
REGION Network 14
   RUNG wire#powerrail
      "FC111_HMI_Status"()
   END_RUNG
   // the same network as SCL:
   "FC111_HMI_Status"();
END_REGION

REGION Network 15
   RUNG wire#powerrail
      "FC500_FAULTS"()
   END_RUNG
   // the same network as SCL:
   "FC500_FAULTS"();
END_REGION

REGION Network 16
   RUNG wire#powerrail
      "FC502_FAULTS C11-C20"()
   END_RUNG
   // the same network as SCL:
   "FC502_FAULTS C11-C20"();
END_REGION

REGION Network 17
   RUNG wire#powerrail
      "FC503_FAULTS C21-C30"()
   END_RUNG
   // the same network as SCL:
   "FC503_FAULTS C21-C30"();
END_REGION

REGION Network 18
   RUNG wire#powerrail
      "FC504_FAULTS C31-C40"()
   END_RUNG
   // the same network as SCL:
   "FC504_FAULTS C31-C40"();
END_REGION

REGION Network 19
   RUNG wire#powerrail
      "FC505_FAULTS C41-C50"()
   END_RUNG
   // the same network as SCL:
   "FC505_FAULTS C41-C50"();
END_REGION

REGION Network 20
   RUNG wire#powerrail
      "FC506_FAULTS C51-C60"()
   END_RUNG
   // the same network as SCL:
   "FC506_FAULTS C51-C60"();
END_REGION

REGION Network 21
   RUNG wire#powerrail
      "FC507_FAULTS C61-C70"()
   END_RUNG
   // the same network as SCL:
   "FC507_FAULTS C61-C70"();
END_REGION

REGION Network 22
   RUNG wire#powerrail
      "FC508_FAULTS C71-C80"()
   END_RUNG
   // the same network as SCL:
   "FC508_FAULTS C71-C80"();
END_REGION

REGION Network 23
   RUNG wire#powerrail
      "FC509_FAULTS C81-C82"()
   END_RUNG
   // the same network as SCL:
   "FC509_FAULTS C81-C82"();
END_REGION

REGION Network 24
   RUNG wire#powerrail
      "FC201_SDC_To_Carrier_Map_IO [C01-C10]"()
   END_RUNG
   // the same network as SCL:
   "FC201_SDC_To_Carrier_Map_IO [C01-C10]"();
END_REGION

REGION Network 25
   RUNG wire#powerrail
      "FC202_SDC_To_Carrier_Map_IO [C11-C20]"()
   END_RUNG
   // the same network as SCL:
   "FC202_SDC_To_Carrier_Map_IO [C11-C20]"();
END_REGION

REGION Network 26
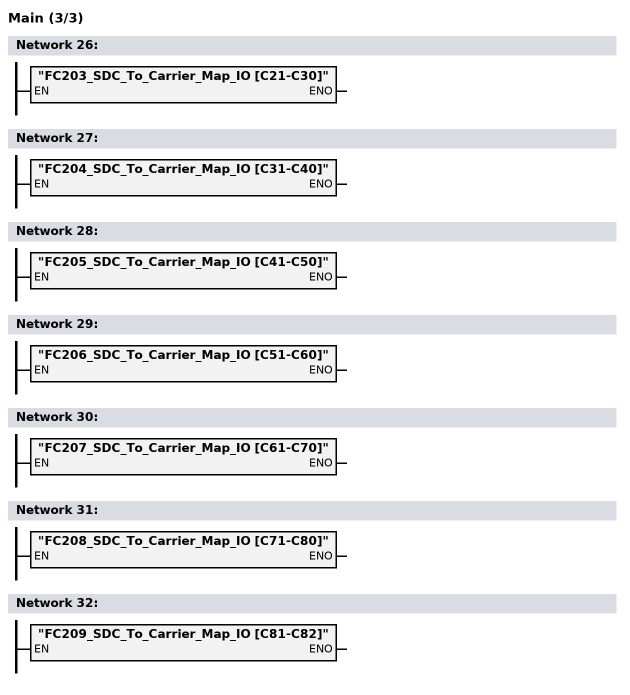
   RUNG wire#powerrail
      "FC203_SDC_To_Carrier_Map_IO [C21-C30]"()
   END_RUNG
   // the same network as SCL:
   "FC203_SDC_To_Carrier_Map_IO [C21-C30]"();
END_REGION

REGION Network 27
   RUNG wire#powerrail
      "FC204_SDC_To_Carrier_Map_IO [C31-C40]"()
   END_RUNG
   // the same network as SCL:
   "FC204_SDC_To_Carrier_Map_IO [C31-C40]"();
END_REGION

REGION Network 28
   RUNG wire#powerrail
      "FC205_SDC_To_Carrier_Map_IO [C41-C50]"()
   END_RUNG
   // the same network as SCL:
   "FC205_SDC_To_Carrier_Map_IO [C41-C50]"();
END_REGION

REGION Network 29
   RUNG wire#powerrail
      "FC206_SDC_To_Carrier_Map_IO [C51-C60]"()
   END_RUNG
   // the same network as SCL:
   "FC206_SDC_To_Carrier_Map_IO [C51-C60]"();
END_REGION

REGION Network 30
   RUNG wire#powerrail
      "FC207_SDC_To_Carrier_Map_IO [C61-C70]"()
   END_RUNG
   // the same network as SCL:
   "FC207_SDC_To_Carrier_Map_IO [C61-C70]"();
END_REGION

REGION Network 31
   RUNG wire#powerrail
      "FC208_SDC_To_Carrier_Map_IO [C71-C80]"()
   END_RUNG
   // the same network as SCL:
   "FC208_SDC_To_Carrier_Map_IO [C71-C80]"();
END_REGION

REGION Network 32
   RUNG wire#powerrail
      "FC209_SDC_To_Carrier_Map_IO [C81-C82]"()
   END_RUNG
   // the same network as SCL:
   "FC209_SDC_To_Carrier_Map_IO [C81-C82]"();
END_REGION
END_ORGANIZATION_BLOCK

ORGANIZATION_BLOCK "Startup"   // OB100, LAD, Startup
TITLE = "Complete Restart"
{ S7_Optimized_Access := 'TRUE' }
VERSION : 0.1
// //============================================================================
// //SIEMENS AG
// //(c)Copyright 2017 All Rights Reserved
// //-----------------------------------------------------------------------------
// //Library: -
// //Tested with: S7-1516-3 PN/DP FW 2.5
// //Engineering: TIA Portal V14 Update1
// //Restrictions: -
// //Requirements: -
// //Functionality: Startup OB for Diagnostics
// //-----------------------------------------------------------------------------
// //Change log table:
// //Version  Date              Expert in charge                               Changes applied
// //01.00.00 25.04.2017 Siemens Industry Online Support First released version
// //============================================================================
   VAR_INPUT
      LostRetentive : Bool;   // True if retentive data are lost
      LostRTC : Bool;   // True if date and time are lost
   END_VAR
   VAR_TEMP
      index : Int;
   END_VAR
BEGIN

REGION Network 1: Set start user diagnostic
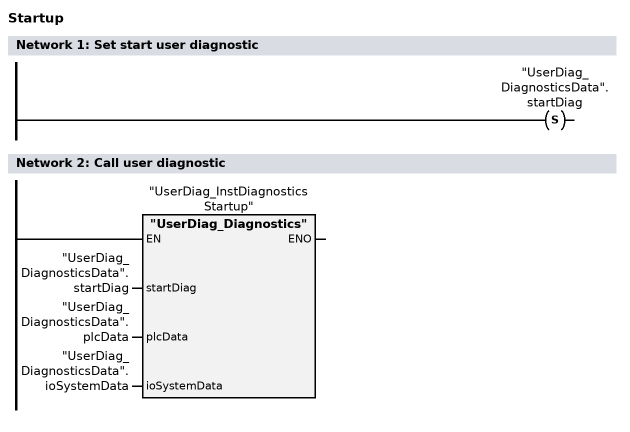
   RUNG wire#powerrail
      S_Coil( "UserDiag_DiagnosticsData".startDiag )
   END_RUNG
   // the same network as SCL:
   "UserDiag_DiagnosticsData".startDiag := TRUE;
END_REGION

REGION Network 2: Call user diagnostic
   RUNG wire#powerrail
      "UserDiag_InstDiagnosticsStartup"(startDiag := "UserDiag_DiagnosticsData".startDiag, plcData := "UserDiag_DiagnosticsData".plcData, ioSystemData := "UserDiag_DiagnosticsData".ioSystemData)
   END_RUNG
   // the same network as SCL:
   "UserDiag_InstDiagnosticsStartup"(startDiag := "UserDiag_DiagnosticsData".startDiag,   // "UserDiag_Diagnostics"
                           plcData := "UserDiag_DiagnosticsData".plcData,
                           ioSystemData := "UserDiag_DiagnosticsData".ioSystemData);
END_REGION
END_ORGANIZATION_BLOCK

ORGANIZATION_BLOCK "Cyclic SDC TO EMS"   // OB300, LAD, CyclicInterrupt
{ S7_Optimized_Access := 'TRUE' }
VERSION : 0.1
   VAR_INPUT
      Initial_Call : Bool;   // Initial call of this OB
      Event_Count : Int;   // Events discarded
   END_VAR
BEGIN
END_ORGANIZATION_BLOCK

// folder: 03_FBs

FUNCTION_BLOCK "FB110_FirstCarrierTCopMotionFB"   // FB110, LAD
{ S7_Optimized_Access := 'TRUE' }
VERSION : 0.1
   VAR_INPUT
      Zone : Int;
      ZonePos : Int;
      ClearOfStopDist : Int;
      StopControlFromEMS01 : "UDT_StopControlFromEMS01";
   END_VAR
   VAR_OUTPUT
      CarrierNumber : Int;
      MoveFwdCommand : Bool;
      DriveCmdSpeed : Int;
      NextCarrierNum : Word;
      NextStopPosition : DWord;
      AtCmdPosition : Bool;
      CarrierInTransitToNextZone : Bool;
      StopStatusToEMS01 : "UDT_StopStatusToEMS01";
   END_VAR
   VAR
      PreviousCarrierNumMemory : Word;
      TrafficCopCarrierZnBuffer : Array[0..40] of "UDT_TrafficCop";
      LastCarrierNextZnPos : Int;
      CarNumZnPos : Int;
      NextZone : Int;
      EndPos_LowLimit : DWord;
      EndPos_HighLimit : DWord;
      ClrOfStopPos_LowLimit : DWord;
      ClrOfStopPos_HighLimit : DWord;
      ClearOfStopPos : DWord;
      ClearToMoveTrain : Bool;
      PrevZone : Int;
      PrevZone_CarrierReady : Bool;
      LastCarrierCurrentZnPos : Int;
      LastCarrierNumber : Word;
      CarrierInTransitToProdZone : Bool;
      ResetCarrierInTransToProd : Bool;
      WaitPositionMemory : DInt;
      OneShot : Bool;
      NextCarrierOffset : DWord;
      PrevZone_EndPos_LowLimit : DWord;
      PrevZone_EndPos_HighLimit : DWord;
   END_VAR
   VAR_TEMP
      NextZoneBuffer : Int;
      LastZone : Int;
      HighSpeedSetpoint : Word;
      LowSpeedSetpoint : Word;
      NextZonePosition : Int;
      NextCarrierOffsetSetup1 : UDInt;
      NextCarrierOffsetSetup2 : UDInt;
   END_VAR
   VAR_TEMP   // added for the SCL form of the ladder/FBD networks
      _w1 : Bool;
      _w2 : Bool;
      _w3 : Bool;
      _w4 : Bool;
      _w5 : Bool;
   END_VAR
BEGIN

REGION Network 1
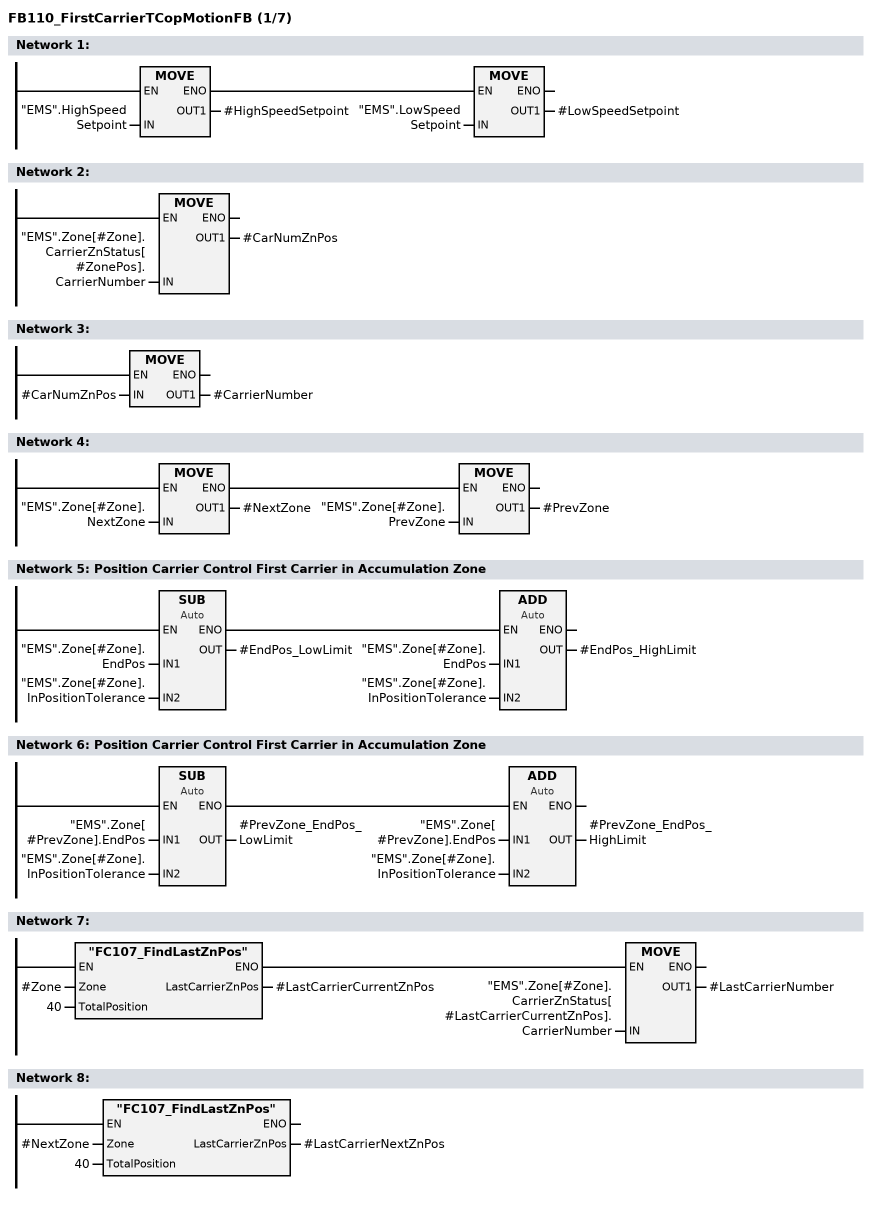
   RUNG wire#powerrail
      Move(in := "EMS".HighSpeedSetpoint, out1 => #HighSpeedSetpoint)
      Move(in := "EMS".LowSpeedSetpoint, out1 => #LowSpeedSetpoint)
   END_RUNG
   // the same network as SCL:
   #HighSpeedSetpoint := "EMS".HighSpeedSetpoint;
   #LowSpeedSetpoint := "EMS".LowSpeedSetpoint;
END_REGION

REGION Network 2
   RUNG wire#powerrail
      Move(in := "EMS".Zone[#Zone].CarrierZnStatus[#ZonePos].CarrierNumber, out1 => #CarNumZnPos)
   END_RUNG
   // the same network as SCL:
   #CarNumZnPos := "EMS".Zone[#Zone].CarrierZnStatus[#ZonePos].CarrierNumber;
END_REGION

REGION Network 3
   RUNG wire#powerrail
      Move(in := #CarNumZnPos, out1 => #CarrierNumber)
   END_RUNG
   // the same network as SCL:
   #CarrierNumber := #CarNumZnPos;
END_REGION

REGION Network 4
   RUNG wire#powerrail
      Move(in := "EMS".Zone[#Zone].NextZone, out1 => #NextZone)
      Move(in := "EMS".Zone[#Zone].PrevZone, out1 => #PrevZone)
   END_RUNG
   // the same network as SCL:
   #NextZone := "EMS".Zone[#Zone].NextZone;
   #PrevZone := "EMS".Zone[#Zone].PrevZone;
END_REGION

REGION Network 5: Position Carrier Control First Carrier in Accumulation Zone
   RUNG wire#powerrail
      Sub(in1 := "EMS".Zone[#Zone].EndPos, in2 := "EMS".Zone[#Zone].InPositionTolerance, out => #EndPos_LowLimit)
      Add(in1 := "EMS".Zone[#Zone].EndPos, in2 := "EMS".Zone[#Zone].InPositionTolerance, out => #EndPos_HighLimit)
   END_RUNG
   // the same network as SCL:
   #EndPos_LowLimit := "EMS".Zone[#Zone].EndPos - "EMS".Zone[#Zone].InPositionTolerance;
   #EndPos_HighLimit := "EMS".Zone[#Zone].EndPos + "EMS".Zone[#Zone].InPositionTolerance;
END_REGION

REGION Network 6: Position Carrier Control First Carrier in Accumulation Zone
   RUNG wire#powerrail
      Sub(in1 := "EMS".Zone[#PrevZone].EndPos, in2 := "EMS".Zone[#Zone].InPositionTolerance, out => #PrevZone_EndPos_LowLimit)
      Add(in1 := "EMS".Zone[#PrevZone].EndPos, in2 := "EMS".Zone[#Zone].InPositionTolerance, out => #PrevZone_EndPos_HighLimit)
   END_RUNG
   // the same network as SCL:
   #PrevZone_EndPos_LowLimit := "EMS".Zone[#PrevZone].EndPos - "EMS".Zone[#Zone].InPositionTolerance;
   #PrevZone_EndPos_HighLimit := "EMS".Zone[#PrevZone].EndPos + "EMS".Zone[#Zone].InPositionTolerance;
END_REGION

REGION Network 7
   RUNG wire#powerrail
      "FC107_FindLastZnPos"(Zone := #Zone, TotalPosition := 40, LastCarrierZnPos => #LastCarrierCurrentZnPos)
      Move(in := "EMS".Zone[#Zone].CarrierZnStatus[#LastCarrierCurrentZnPos].CarrierNumber, out1 => #LastCarrierNumber)
   END_RUNG
   // the same network as SCL:
   "FC107_FindLastZnPos"(Zone := #Zone,
                         TotalPosition := 40,
                         LastCarrierZnPos => #LastCarrierCurrentZnPos,
                         ENO => #_w1);
   IF #_w1 THEN
       #LastCarrierNumber := "EMS".Zone[#Zone].CarrierZnStatus[#LastCarrierCurrentZnPos].CarrierNumber;
   END_IF;
END_REGION

REGION Network 8
   RUNG wire#powerrail
      "FC107_FindLastZnPos"(Zone := #NextZone, TotalPosition := 40, LastCarrierZnPos => #LastCarrierNextZnPos)
   END_RUNG
   // the same network as SCL:
   "FC107_FindLastZnPos"(Zone := #NextZone, TotalPosition := 40, LastCarrierZnPos => #LastCarrierNextZnPos);
END_REGION

REGION Network 9: Position Carrier Control First Carrier in Production Zone
   // Control of First Carrier in Zone Closest to end position/Stop.  Move command is issued to carrier. Carrier will move in auto.
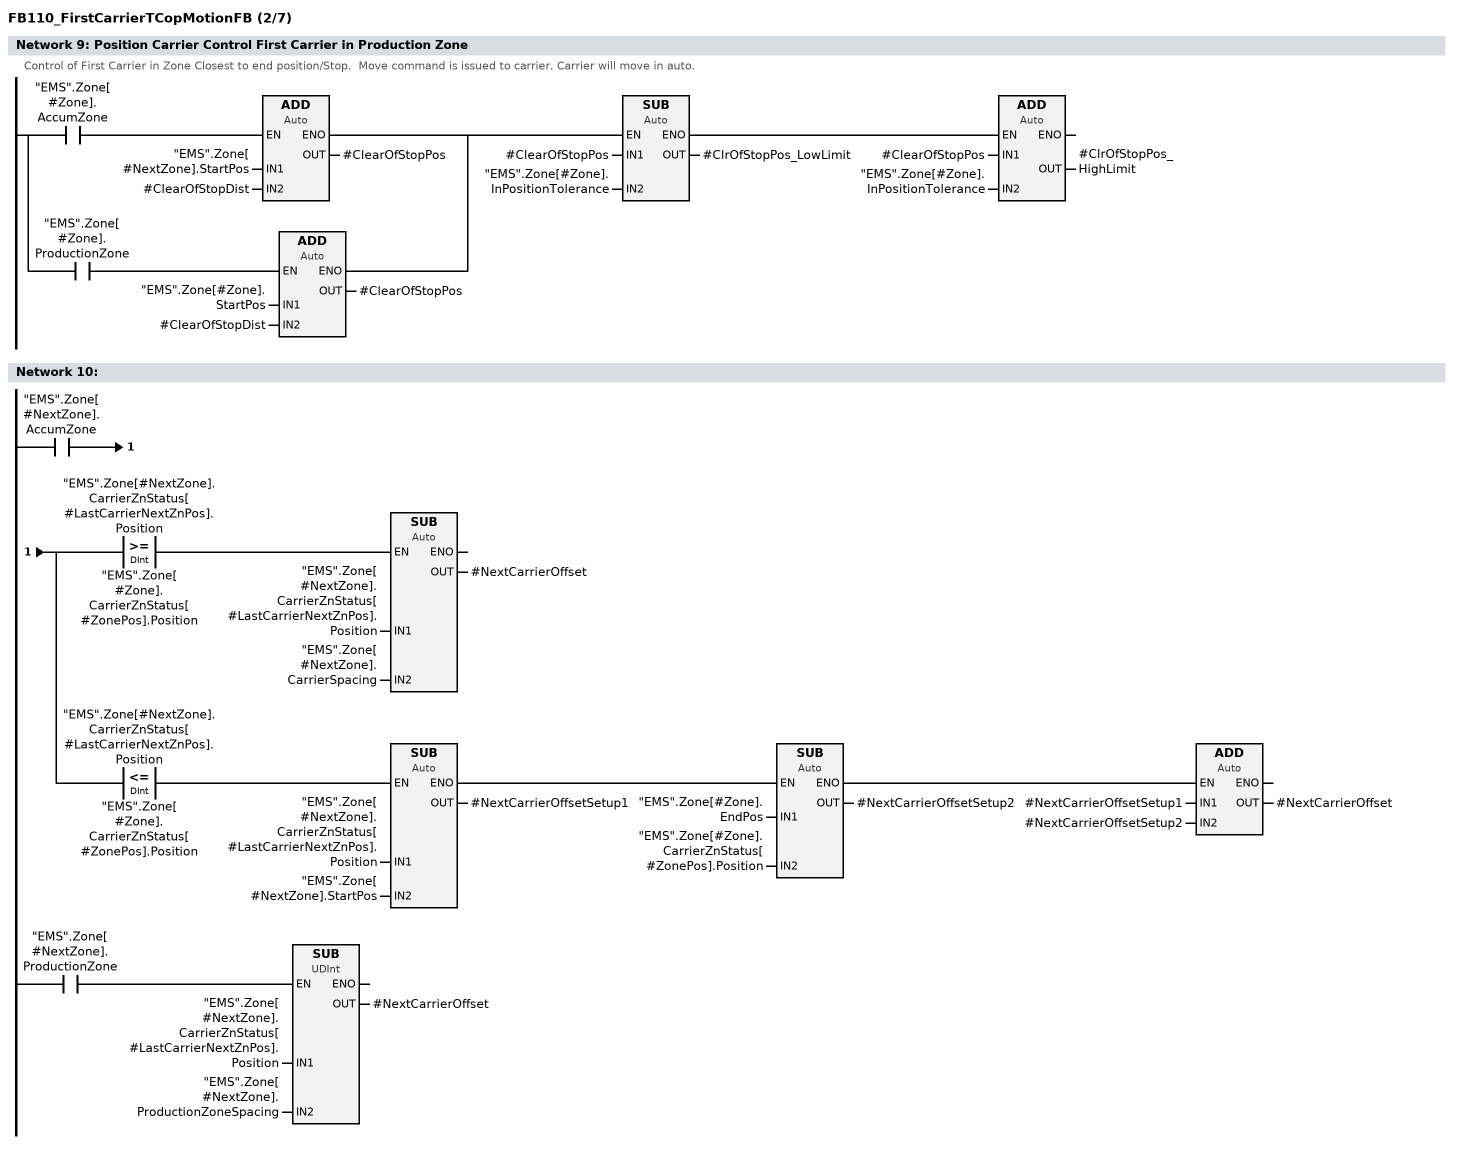
   RUNG wire#powerrail
      Contact( "EMS".Zone[#Zone].AccumZone )
      Add(in1 := "EMS".Zone[#NextZone].StartPos, in2 := #ClearOfStopDist, out => #ClearOfStopPos)
      wire#w1
      Sub(in1 := #ClearOfStopPos, in2 := "EMS".Zone[#Zone].InPositionTolerance, out => #ClrOfStopPos_LowLimit)
      Add(in1 := #ClearOfStopPos, in2 := "EMS".Zone[#Zone].InPositionTolerance, out => #ClrOfStopPos_HighLimit)
   END_RUNG
   RUNG wire#powerrail
      Contact( "EMS".Zone[#Zone].ProductionZone )
      Add(in1 := "EMS".Zone[#Zone].StartPos, in2 := #ClearOfStopDist, out => #ClearOfStopPos)
   END_RUNG wire#w1
   // the same network as SCL:
   IF "EMS".Zone[#Zone].AccumZone THEN
       #ClearOfStopPos := "EMS".Zone[#NextZone].StartPos + #ClearOfStopDist;
   END_IF;
   IF "EMS".Zone[#Zone].ProductionZone THEN
       #ClearOfStopPos := "EMS".Zone[#Zone].StartPos + #ClearOfStopDist;
   END_IF;
   IF "EMS".Zone[#Zone].AccumZone OR "EMS".Zone[#Zone].ProductionZone THEN
       #ClrOfStopPos_LowLimit := #ClearOfStopPos - "EMS".Zone[#Zone].InPositionTolerance;
       #ClrOfStopPos_HighLimit := #ClearOfStopPos + "EMS".Zone[#Zone].InPositionTolerance;
   END_IF;
END_REGION

REGION Network 10
   RUNG wire#powerrail
      Contact( "EMS".Zone[#NextZone].AccumZone )
      wire#w1
      { S7_Templates := "SrcType := DInt" } GE_Contact(in1 := "EMS".Zone[#NextZone].CarrierZnStatus[#LastCarrierNextZnPos].Position, in2 := "EMS".Zone[#Zone].CarrierZnStatus[#ZonePos].Position)
      Sub(in1 := "EMS".Zone[#NextZone].CarrierZnStatus[#LastCarrierNextZnPos].Position, in2 := "EMS".Zone[#NextZone].CarrierSpacing, out => #NextCarrierOffset)
   END_RUNG
   RUNG wire#w1
      { S7_Templates := "SrcType := DInt" } LE_Contact(in1 := "EMS".Zone[#NextZone].CarrierZnStatus[#LastCarrierNextZnPos].Position, in2 := "EMS".Zone[#Zone].CarrierZnStatus[#ZonePos].Position)
      Sub(in1 := "EMS".Zone[#NextZone].CarrierZnStatus[#LastCarrierNextZnPos].Position, in2 := "EMS".Zone[#NextZone].StartPos, out => #NextCarrierOffsetSetup1)
      Sub(in1 := "EMS".Zone[#Zone].EndPos, in2 := "EMS".Zone[#Zone].CarrierZnStatus[#ZonePos].Position, out => #NextCarrierOffsetSetup2)
      Add(in1 := #NextCarrierOffsetSetup1, in2 := #NextCarrierOffsetSetup2, out => #NextCarrierOffset)
   END_RUNG
   RUNG wire#powerrail
      Contact( "EMS".Zone[#NextZone].ProductionZone )
      { S7_Templates := "SrcType := UDInt" } Sub(in1 := "EMS".Zone[#NextZone].CarrierZnStatus[#LastCarrierNextZnPos].Position, in2 := "EMS".Zone[#NextZone].ProductionZoneSpacing, out => #NextCarrierOffset)
   END_RUNG
   // the same network as SCL:
   IF "EMS".Zone[#NextZone].AccumZone AND ("EMS".Zone[#NextZone].CarrierZnStatus[#LastCarrierNextZnPos].Position >= "EMS".Zone[#Zone].CarrierZnStatus[#ZonePos].Position) THEN
       #NextCarrierOffset := "EMS".Zone[#NextZone].CarrierZnStatus[#LastCarrierNextZnPos].Position - "EMS".Zone[#NextZone].CarrierSpacing;
   END_IF;
   IF "EMS".Zone[#NextZone].AccumZone AND ("EMS".Zone[#NextZone].CarrierZnStatus[#LastCarrierNextZnPos].Position <= "EMS".Zone[#Zone].CarrierZnStatus[#ZonePos].Position) THEN
       #NextCarrierOffsetSetup1 := "EMS".Zone[#NextZone].CarrierZnStatus[#LastCarrierNextZnPos].Position - "EMS".Zone[#NextZone].StartPos;
       #NextCarrierOffsetSetup2 := "EMS".Zone[#Zone].EndPos - "EMS".Zone[#Zone].CarrierZnStatus[#ZonePos].Position;
       #NextCarrierOffset := #NextCarrierOffsetSetup1 + #NextCarrierOffsetSetup2;
   END_IF;
   IF "EMS".Zone[#NextZone].ProductionZone THEN
       #NextCarrierOffset := "EMS".Zone[#NextZone].CarrierZnStatus[#LastCarrierNextZnPos].Position - "EMS".Zone[#NextZone].ProductionZoneSpacing;
   END_IF;
END_REGION

REGION Network 11
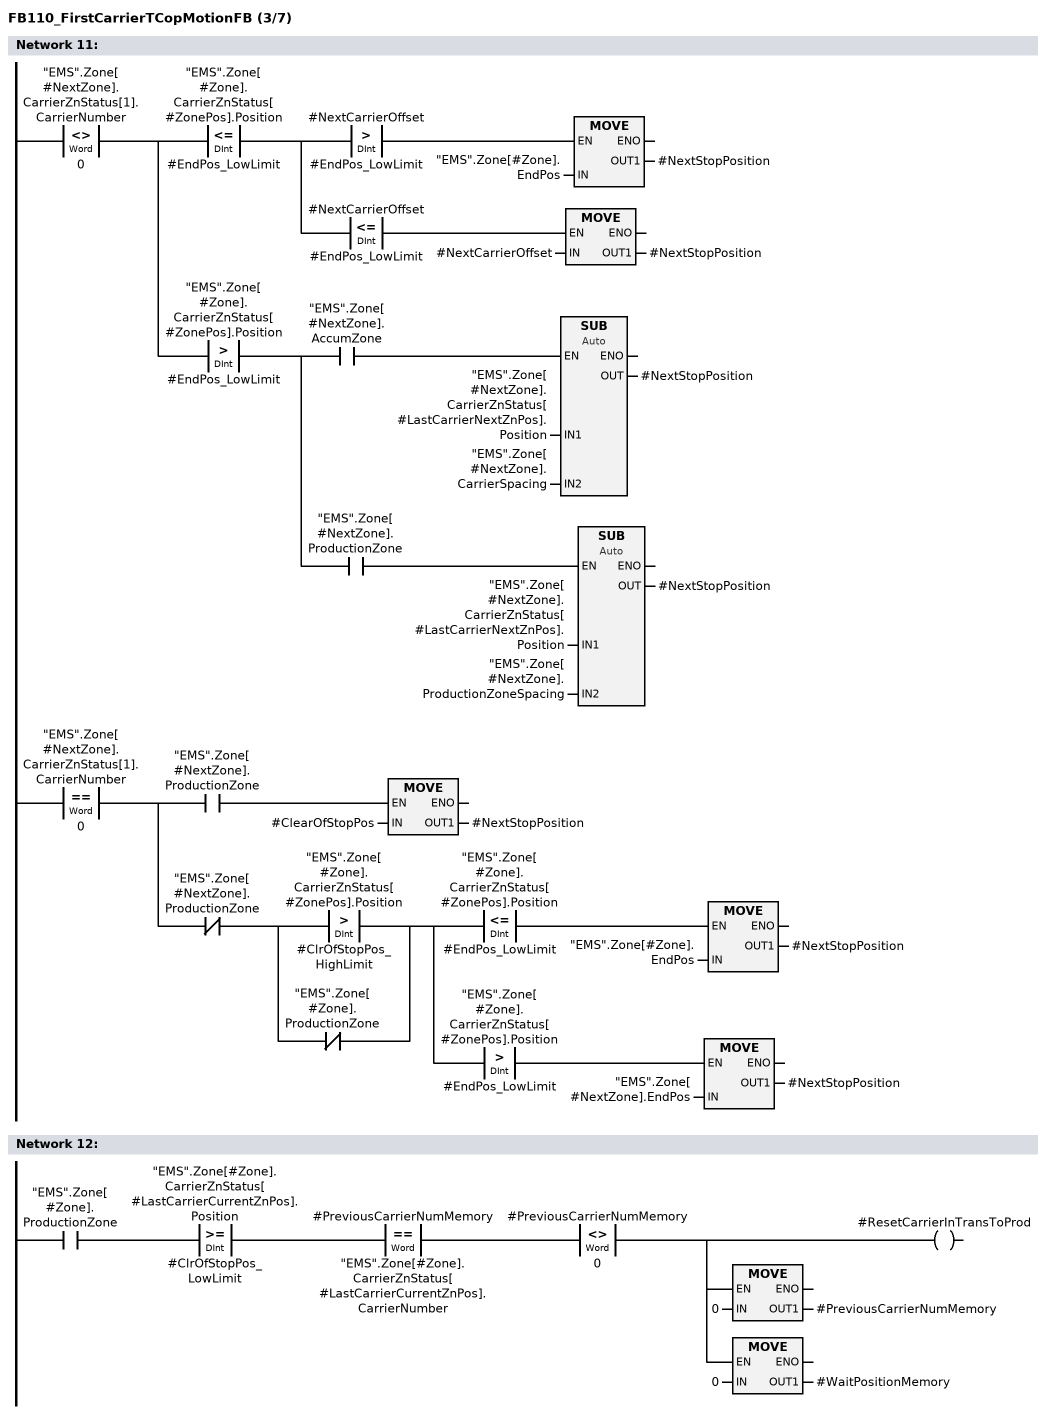
   RUNG wire#powerrail
      { S7_Templates := "SrcType := Word" } NE_Contact(in1 := "EMS".Zone[#NextZone].CarrierZnStatus[1].CarrierNumber, in2 := 0)
      wire#w1
      { S7_Templates := "SrcType := DInt" } LE_Contact(in1 := "EMS".Zone[#Zone].CarrierZnStatus[#ZonePos].Position, in2 := #EndPos_LowLimit)
      wire#w2
      { S7_Templates := "SrcType := DInt" } GT_Contact(in1 := #NextCarrierOffset, in2 := #EndPos_LowLimit)
      Move(in := "EMS".Zone[#Zone].EndPos, out1 => #NextStopPosition)
   END_RUNG
   RUNG wire#w2
      { S7_Templates := "SrcType := DInt" } LE_Contact(in1 := #NextCarrierOffset, in2 := #EndPos_LowLimit)
      Move(in := #NextCarrierOffset, out1 => #NextStopPosition)
   END_RUNG
   RUNG wire#w1
      { S7_Templates := "SrcType := DInt" } GT_Contact(in1 := "EMS".Zone[#Zone].CarrierZnStatus[#ZonePos].Position, in2 := #EndPos_LowLimit)
      wire#w3
      Contact( "EMS".Zone[#NextZone].AccumZone )
      Sub(in1 := "EMS".Zone[#NextZone].CarrierZnStatus[#LastCarrierNextZnPos].Position, in2 := "EMS".Zone[#NextZone].CarrierSpacing, out => #NextStopPosition)
   END_RUNG
   RUNG wire#w3
      Contact( "EMS".Zone[#NextZone].ProductionZone )
      Sub(in1 := "EMS".Zone[#NextZone].CarrierZnStatus[#LastCarrierNextZnPos].Position, in2 := "EMS".Zone[#NextZone].ProductionZoneSpacing, out => #NextStopPosition)
   END_RUNG
   RUNG wire#powerrail
      { S7_Templates := "SrcType := Word" } EQ_Contact(in1 := "EMS".Zone[#NextZone].CarrierZnStatus[1].CarrierNumber, in2 := 0)
      wire#w4
      Contact( "EMS".Zone[#NextZone].ProductionZone )
      Move(in := #ClearOfStopPos, out1 => #NextStopPosition)
   END_RUNG
   RUNG wire#w4
      I_Contact( "EMS".Zone[#NextZone].ProductionZone )
      wire#w5
      { S7_Templates := "SrcType := DInt" } GT_Contact(in1 := "EMS".Zone[#Zone].CarrierZnStatus[#ZonePos].Position, in2 := #ClrOfStopPos_HighLimit)
      wire#w6
      { S7_Templates := "SrcType := DInt" } LE_Contact(in1 := "EMS".Zone[#Zone].CarrierZnStatus[#ZonePos].Position, in2 := #EndPos_LowLimit)
      Move(in := "EMS".Zone[#Zone].EndPos, out1 => #NextStopPosition)
   END_RUNG
   RUNG wire#w5
      I_Contact( "EMS".Zone[#Zone].ProductionZone )
   END_RUNG wire#w6
   RUNG wire#w6
      { S7_Templates := "SrcType := DInt" } GT_Contact(in1 := "EMS".Zone[#Zone].CarrierZnStatus[#ZonePos].Position, in2 := #EndPos_LowLimit)
      Move(in := "EMS".Zone[#NextZone].EndPos, out1 => #NextStopPosition)
   END_RUNG
   // the same network as SCL:
   #_w1 := "EMS".Zone[#NextZone].CarrierZnStatus[1].CarrierNumber <> 0;
   #_w2 := #_w1 AND ("EMS".Zone[#Zone].CarrierZnStatus[#ZonePos].Position <= #EndPos_LowLimit);
   IF #_w2 AND (#NextCarrierOffset > #EndPos_LowLimit) THEN
       #NextStopPosition := "EMS".Zone[#Zone].EndPos;
   END_IF;
   IF #_w2 AND (#NextCarrierOffset <= #EndPos_LowLimit) THEN #NextStopPosition := #NextCarrierOffset; END_IF;
   #_w3 := #_w1 AND ("EMS".Zone[#Zone].CarrierZnStatus[#ZonePos].Position > #EndPos_LowLimit);
   IF #_w3 AND "EMS".Zone[#NextZone].AccumZone THEN
       #NextStopPosition := "EMS".Zone[#NextZone].CarrierZnStatus[#LastCarrierNextZnPos].Position - "EMS".Zone[#NextZone].CarrierSpacing;
   END_IF;
   IF #_w3 AND "EMS".Zone[#NextZone].ProductionZone THEN
       #NextStopPosition := "EMS".Zone[#NextZone].CarrierZnStatus[#LastCarrierNextZnPos].Position - "EMS".Zone[#NextZone].ProductionZoneSpacing;
   END_IF;
   #_w4 := "EMS".Zone[#NextZone].CarrierZnStatus[1].CarrierNumber = 0;
   IF #_w4 AND "EMS".Zone[#NextZone].ProductionZone THEN #NextStopPosition := #ClearOfStopPos; END_IF;
   #_w5 := #_w4 AND NOT "EMS".Zone[#NextZone].ProductionZone AND (("EMS".Zone[#Zone].CarrierZnStatus[#ZonePos].Position > #ClrOfStopPos_HighLimit) OR NOT "EMS".Zone[#Zone].ProductionZone);
   IF #_w5 AND ("EMS".Zone[#Zone].CarrierZnStatus[#ZonePos].Position <= #EndPos_LowLimit) THEN
       #NextStopPosition := "EMS".Zone[#Zone].EndPos;
   END_IF;
   IF #_w5 AND ("EMS".Zone[#Zone].CarrierZnStatus[#ZonePos].Position > #EndPos_LowLimit) THEN
       #NextStopPosition := "EMS".Zone[#NextZone].EndPos;
   END_IF;
END_REGION

REGION Network 12
   RUNG wire#powerrail
      Contact( "EMS".Zone[#Zone].ProductionZone )
      { S7_Templates := "SrcType := DInt" } GE_Contact(in1 := "EMS".Zone[#Zone].CarrierZnStatus[#LastCarrierCurrentZnPos].Position, in2 := #ClrOfStopPos_LowLimit)
      { S7_Templates := "SrcType := Word" } EQ_Contact(in1 := #PreviousCarrierNumMemory, in2 := "EMS".Zone[#Zone].CarrierZnStatus[#LastCarrierCurrentZnPos].CarrierNumber)
      { S7_Templates := "SrcType := Word" } NE_Contact(in1 := #PreviousCarrierNumMemory, in2 := 0)
      wire#w1
      Coil( #ResetCarrierInTransToProd )
   END_RUNG
   RUNG wire#w1
      Move(in := 0, out1 => #PreviousCarrierNumMemory)
   END_RUNG
   RUNG wire#w1
      Move(in := 0, out1 => #WaitPositionMemory)
   END_RUNG
   // the same network as SCL:
   #ResetCarrierInTransToProd := "EMS".Zone[#Zone].ProductionZone AND ("EMS".Zone[#Zone].CarrierZnStatus[#LastCarrierCurrentZnPos].Position >= #ClrOfStopPos_LowLimit) AND (#PreviousCarrierNumMemory = "EMS".Zone[#Zone].CarrierZnStatus[#LastCarrierCurrentZnPos].CarrierNumber) AND (#PreviousCarrierNumMemory <> 0);
   IF #ResetCarrierInTransToProd THEN
       #PreviousCarrierNumMemory := 0;
       #WaitPositionMemory := 0;
   END_IF;
END_REGION

REGION Network 13
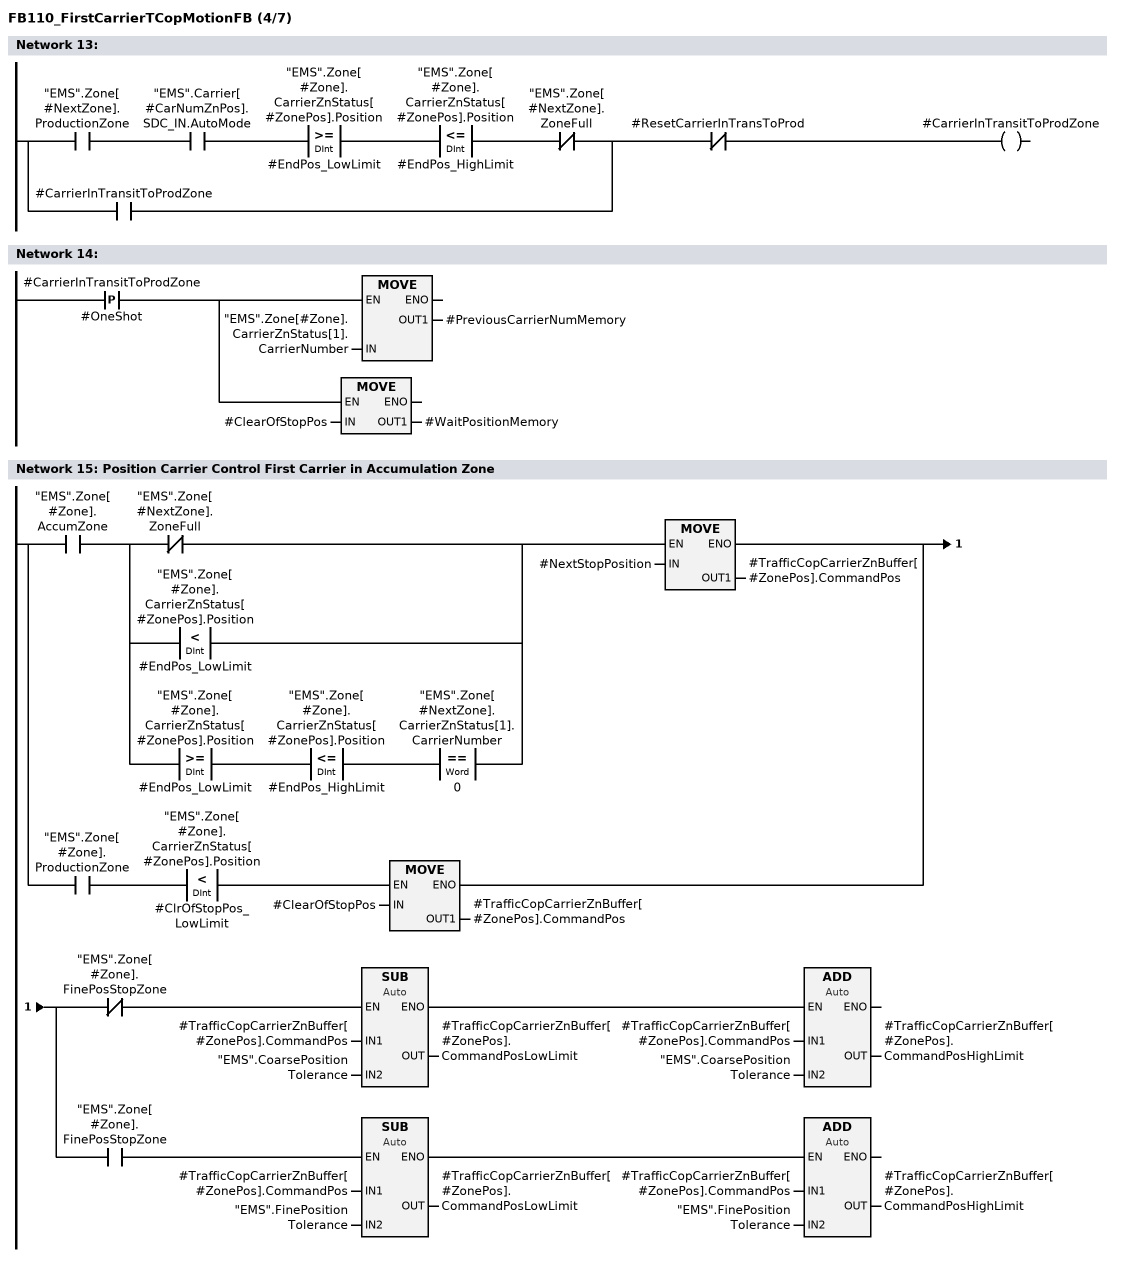
   RUNG wire#powerrail
      Contact( "EMS".Zone[#NextZone].ProductionZone )
      Contact( "EMS".Carrier[#CarNumZnPos].SDC_IN.AutoMode )
      { S7_Templates := "SrcType := DInt" } GE_Contact(in1 := "EMS".Zone[#Zone].CarrierZnStatus[#ZonePos].Position, in2 := #EndPos_LowLimit)
      { S7_Templates := "SrcType := DInt" } LE_Contact(in1 := "EMS".Zone[#Zone].CarrierZnStatus[#ZonePos].Position, in2 := #EndPos_HighLimit)
      I_Contact( "EMS".Zone[#NextZone].ZoneFull )
      wire#w1
      I_Contact( #ResetCarrierInTransToProd )
      Coil( #CarrierInTransitToProdZone )
   END_RUNG
   RUNG wire#powerrail
      Contact( #CarrierInTransitToProdZone )
   END_RUNG wire#w1
   // the same network as SCL:
   #CarrierInTransitToProdZone := (("EMS".Zone[#NextZone].ProductionZone AND "EMS".Carrier[#CarNumZnPos].SDC_IN.AutoMode AND ("EMS".Zone[#Zone].CarrierZnStatus[#ZonePos].Position >= #EndPos_LowLimit) AND ("EMS".Zone[#Zone].CarrierZnStatus[#ZonePos].Position <= #EndPos_HighLimit) AND NOT "EMS".Zone[#NextZone].ZoneFull) OR #CarrierInTransitToProdZone) AND NOT #ResetCarrierInTransToProd;
END_REGION

REGION Network 14
   RUNG wire#powerrail
      P_Contact(operand := #CarrierInTransitToProdZone, bit := #OneShot)
      wire#w1
      Move(in := "EMS".Zone[#Zone].CarrierZnStatus[1].CarrierNumber, out1 => #PreviousCarrierNumMemory)
   END_RUNG
   RUNG wire#w1
      Move(in := #ClearOfStopPos, out1 => #WaitPositionMemory)
   END_RUNG
   // the same network as SCL:
   #_w1 := #CarrierInTransitToProdZone AND NOT #OneShot;   // rising edge of #CarrierInTransitToProdZone
   #OneShot := #CarrierInTransitToProdZone;
   IF #_w1 THEN
       #PreviousCarrierNumMemory := "EMS".Zone[#Zone].CarrierZnStatus[1].CarrierNumber;
       #WaitPositionMemory := #ClearOfStopPos;
   END_IF;
END_REGION
